        [25]   // Subsurface Cutter Alarm Tone Generation Counter
        [11]   // TRIM DECK Fault Tracking: Number of Times M2CM12N Drive Faulted
        [12]   // TRIM DECK Fault Tracking: Number of Times M2CM04N Drive Faulted
        [18]   // TRIM DECK Fault Tracking: Number of Times M2CM10S Drive Faulted
        [1]   // TRIM DECK Fault Tracking: Number of Times M2CM02 Drive Faulted
        [19]   // TRIM DECK Fault Tracking: Number of Times M2CM11S Drive Faulted
        [22]   // Debug Counter Number of Times M2CM09 Drive Faulted
        [23]   // Debug Counter Number of Times M2CM10 Drive Faulted
        [30]   // TRIM DECK Fault Tracking: Number of Times M2CM01 Drive is Stopped
   C50 : COUNTER[33];
        [10]   // Conveyor 10 Phantom Caps Generated Counter
        [11]   // Conveyor 11 Phantom Caps Generated Counter
        [12]   // Conveyor 12 Phantom Caps Generated Counter
        [13]   // Conveyor 13 Phantom Caps Generated Counter
        [14]   // Conveyor 14 Phantom Caps Generated Counter
        [15]   // Conveyor 15 Phantom Caps Generated Counter
        [16]   // Conveyor 16 Phantom Caps Generated Counter
        [17]   // Conveyor 17 Phantom Caps Generated Counter
        [18]   // Conveyor 18 Phantom Caps Generated Counter
        [19]   // Conveyor 19 Phantom Caps Generated Counter
        [1]   // Conveyor 1 Phantom Caps Generated Counter
        [20]   // Conveyor 20 Phantom Caps Generated Counter
        [21]   // Conveyor 21 Phantom Caps Generated Counter
        [22]   // Conveyor 22 Phantom Caps Generated Counter
        [23]   // Conveyor 23 Phantom Caps Generated Counter
        [24]   // Conveyor 24 Phantom Caps Generated Counter
        [25]   // Conveyor 25 Phantom Caps Generated Counter
        [26]   // Conveyor 26 Phantom Caps Generated Counter
        [27]   // Conveyor 27 Phantom Caps Generated Counter
        [28]   // Conveyor 28 Phantom Caps Generated Counter
        [29]   // Conveyor 29 Phantom Caps Generated Counter
        [2]   // Conveyor 2 Phantom Caps Generated Counter
        [30]   // Conveyor 30 Phantom Caps Generated Counter
        [31]   // Conveyor 31 Phantom Caps Generated Counter
        [32]   // Conveyor 32 Phantom Caps Generated Counter
        [3]   // Conveyor 3 Phantom Caps Generated Counter
        [4]   // Conveyor 4 Phantom Caps Generated Counter
        [5]   // Conveyor 5 Phantom Caps Generated Counter
        [6]   // Conveyor 6 Phantom Caps Generated Counter
        [7]   // Conveyor 7 Phantom Caps Generated Counter
        [8]   // Conveyor 8 Phantom Caps Generated Counter
        [9]   // Conveyor 9 Phantom Caps Generated Counter
   C61 : COUNTER[33];
        [5]   // Conveyor 5 Glass in Transit Counter
        [6]   // Conveyor 6 Glass in Transit Counter
        [7]   // Conveyor 7 Glass in Transit Counter
        [8]   // Conveyor 8 Glass in Transit Counter
        [9]   // Conveyor 9 Glass in Transit Counter
        [17]   // Conveyor 17 Glass in Transit Counter
        [18]   // Conveyor 18 Glass in Transit Counter
        [19]   // Conveyor 19 Glass in Transit Counter
        [1]   // Conveyor 1 Glass in Transit Counter
        [20]   // Conveyor 20 Glass in Transit Counter
        [21]   // Conveyor 21 Glass in Transit Counter
        [22]   // Conveyor 22 Glass in Transit Counter
        [23]   // Conveyor 23 Glass in Transit Counter
        [24]   // Conveyor 24 Glass in Transit Counter
        [25]   // Conveyor 25 Glass in Transit Counter
        [26]   // Conveyor 26 Glass in Transit Counter
        [27]   // Conveyor 27 Glass in Transit Counter
        [10]   // Conveyor 10 Glass in Transit Counter
        [11]   // Conveyor 11 Glass in Transit Counter
        [12]   // Conveyor 12 Glass in Transit Counter
        [13]   // Conveyor 13 Glass in Transit Counter
        [14]   // Conveyor 14 Glass in Transit Counter
        [15]   // Conveyor 15 Glass in Transit Counter
        [28]   // Conveyor 28 Glass in Transit Counter
        [29]   // Conveyor 29 Glass in Transit Counter
        [2]   // Conveyor 2 Glass in Transit Counter
        [16]   // Conveyor 16 Glass in Transit Counter
        [30]   // Conveyor 30 Glass in Transit Counter
        [31]   // Conveyor 31 Glass in Transit Counter
        [32]   // Conveyor 32 Glass in Transit Counter
        [3]   // Conveyor 3 Glass in Transit Counter
        [4]   // Conveyor 4 Glass in Transit Counter
   CM_AreaStackerToLine_JS1 : CM_AreaStackerToLine; {access Read Only}
   CM_AreaStackerToLine_JS1_Sync : CM_AreaStackerToLine := (dSyncHead := 612195157, xAreaOk := 1, xStackerInUnloaderMode := 1, iPresetNumberPlateOnRack[0] := 30, iPresetNumberPlateOnRack[1] := 30, iActualNumberPlateOnRack[0] := 24, iActualNumberPlateOnRack[1] := 23, dGap_cmm := 25000, dMsgDataSyncFdbk := 230589, dMsgDataSync := 289, dMsgOPTSyncFdbk := 339568305, dMsgOPTSync := 297768899, dSyncTail := 612195157);
        .iPresetNumberPlateOnRack[0]   // RHS
        .iActualNumberPlateOnRack[0]   // RHS
        .iActualNumberPlateOnRack[1]   // LHS
        .iPresetNumberPlateOnRack[1]   // LHS
        .dGap_cmm   // [mm/100]
   CM_AreaStackerToLine_JS2 : CM_AreaStackerToLine; {access Read Only}
   CM_AreaStackerToLine_JS2_Sync : CM_AreaStackerToLine := (dSyncHead := 612195157, xAreaOk := 1, xStackerInUnloaderMode := 1, iPresetNumberPlateOnRack[0] := 30, iPresetNumberPlateOnRack[1] := 30, iActualNumberPlateOnRack[0] := 24, iActualNumberPlateOnRack[1] := 23, dGap_cmm := 25000, dMsgDataSyncFdbk := 230589, dMsgDataSync := 289, dMsgOPTSyncFdbk := 339568305, dMsgOPTSync := 297768899, dSyncTail := 612195157);
        .iPresetNumberPlateOnRack[0]   // RHS
        .iPresetNumberPlateOnRack[1]   // LHS
        .iActualNumberPlateOnRack[0]   // RHS
        .iActualNumberPlateOnRack[1]   // LHS
        .dGap_cmm   // [mm/100]
   CM_ConveyorStackerToLine_JS1 : CM_ConveyorStackerToLine; {access Read Only}
   CM_ConveyorStackerToLine_JS1_Sync : CM_ConveyorStackerToLine := (dSyncHead := 598734532, xCycleOn := 1, xConditionOkForStopCycle := 1, xInitialContionOk := 1, xOutputEnable := 1, xAirMode := 1, dSyncTail := 598734532);
   CM_ConveyorStackerToLine_JS2 : CM_ConveyorStackerToLine; {access Read Only}
   CM_ConveyorStackerToLine_JS2_Sync : CM_ConveyorStackerToLine := (dSyncHead := 598734532, xCycleOn := 1, xConditionOkForStopCycle := 1, xInitialContionOk := 1, xOutputEnable := 1, xAirMode := 1, dSyncTail := 598734532);
   CM_DATA_Snap_Rx : CM_DATA_Z200; {access Read Only}
   CM_DATA_Snap_Rx_TempBuffer : SINT[696]; {access Read Only}
   CM_DATA_Z410_Rx : UDT_PlateData_Convoy; {access Read Only}
   CM_DATA_Z410_Rx_Sync : UDT_PlateData_Convoy; {access Read Only}
   CM_DATA_Z410_Rx_TmpBuffer : SINT[104]; {access Read Only}
   CM_DATA_Z410_Tx : UDT_PlateData_Convoy; {access Read Only}
   CM_DATA_Z410_Tx_MSG : MESSAGE; {access Read Only}
   CM_DATA_Z410_Tx_PH : DINT; {access Read Only}
   CM_DATA_Z410_Tx_TempBuffer : SINT[104]; {access Read Only}
   CM_DATA_Z410_Tx_tmON : TIMER; {access Read Only}
   CM_DATA_Z420_Rx : UDT_PlateData_Convoy; {access Read Only}
   CM_DATA_Z420_Rx_Sync : UDT_PlateData_Convoy; {access Read Only}
   CM_DATA_Z420_Rx_TmpBuffer : SINT[104]; {access Read Only}
   CM_DATA_Z420_Tx : UDT_PlateData_Convoy; {access Read Only}
   CM_DATA_Z420_Tx_MSG : MESSAGE; {access Read Only}
   CM_DATA_Z420_Tx_PH : DINT; {access Read Only}
   CM_DATA_Z420_Tx_TempBuffer : SINT[104]; {access Read Only}
   CM_DATA_Z420_Tx_tmON : TIMER; {access Read Only}
   CM_INPUT_Z200 : CM_INPUT_Z200; {access Read Only}
   CM_INPUT_Z200_Sync : CM_INPUT_Z200; {access Read Only}
   CM_LineToAreaStacker_JS1 : CM_LineToAreaStacker := (dSyncHead := 612195196, xConditionOkForAccessArea := 1, dMsgDataSyncFdbk := 289, dMsgDataSync := 230589, dMsgOPTSyncFdbk := 297768899, dMsgOPTSync := 339568321, dSyncTail := 612195196); {produced}
   CM_LineToAreaStacker_JS2 : CM_LineToAreaStacker := (dSyncHead := 612195196, xConditionOkForAccessArea := 1, dMsgDataSyncFdbk := 289, dMsgDataSync := 230589, dMsgOPTSyncFdbk := 297768899, dMsgOPTSync := 339568321, dSyncTail := 612195196); {produced}
   CM_LineToConveyorStacker_JS1 : CM_LineToConveyorStacker := (dSyncHead := 598734505, xEmergencyOn := 1, xLineCycleOn := 1, xOutputEnable := 1, xReadyToMove := 1, dLineSpeed_dmm_min := 600000, dSyncTail := 598734505); {produced}
   CM_LineToConveyorStacker_JS2 : CM_LineToConveyorStacker := (dSyncHead := 598734505, xEmergencyOn := 1, xLineCycleOn := 1, xOutputEnable := 1, xReadyToMove := 1, dLineSpeed_dmm_min := 600000, dSyncTail := 598734505); {produced}
   CM_OUTPUT_Z200 : CM_OUTPUT_Z200; {access Read Only}
   CNV10_COP_BUFR : ALIAS FOR N31[10];
   CNV10_FLT : ALIAS FOR I[4].9;
   CNV10_FWD : ALIAS FOR O[5].9;
   CNV10_LENGTH : ALIAS FOR N32[10];
   CNV10_LOST : ALIAS FOR C48[10];
   CNV10_PHNTM : ALIAS FOR C50[10];
   CNV10_RES_CAPID : ALIAS FOR N40[10];
   CNV10_RESIN : ALIAS FOR B42[0].10;
   CNV10_RESIN_DEB : ALIAS FOR T47[10];
   CNV10_RESIN_LED : ALIAS FOR B45[0].10;
   CNV10_RESIN_TR : ALIAS FOR B46[0].10;
   CNV10_RESOUT : ALIAS FOR B43[0].10;
   CNV10_REV : ALIAS FOR O[6].9;
   CNV10_RTUNE : ALIAS FOR C49[10];
   CNV10_SS1 : ALIAS FOR O[8].9;
   CNV10_SS2 : ALIAS FOR O[7].9;
   CNV10_T : ALIAS FOR B60[0].10;
   CNV10_T_CNTRS : ALIAS FOR C61[10];
   CNV10_WIN : ALIAS FOR B41[0].10;
   CNV11_COP_BUFR : ALIAS FOR N31[11];
   CNV11_FLT : ALIAS FOR I[4].10;
   CNV11_FWD : ALIAS FOR O[5].10;
   CNV11_LENGTH : ALIAS FOR N32[11];
   CNV11_LOST : ALIAS FOR C48[11];
   CNV11_PHNTM : ALIAS FOR C50[11];
   CNV11_RES_CAPID : ALIAS FOR N40[11];
   CNV11_RESIN : ALIAS FOR B42[0].11;
   CNV11_RESIN_DEB : ALIAS FOR T47[11];
   CNV11_RESIN_LED : ALIAS FOR B45[0].11;
   CNV11_RESIN_TR : ALIAS FOR B46[0].11;
   CNV11_RESOUT : ALIAS FOR B43[0].11;
   CNV11_REV : ALIAS FOR O[6].10;
   CNV11_RTUNE : ALIAS FOR C49[11];
   CNV11_SS1 : ALIAS FOR O[8].10;
   CNV11_SS2 : ALIAS FOR O[7].10;
   CNV11_T : ALIAS FOR B60[0].11;
   CNV11_T_CNTRS : ALIAS FOR C61[11];
   CNV11_WIN : ALIAS FOR B41[0].11;
   CNV12_COP_BUFR : ALIAS FOR N31[12];
   CNV12_FLT : ALIAS FOR I[4].11;
   CNV12_LENGTH : ALIAS FOR N32[12];
   CNV12_LOST : ALIAS FOR C48[12];
   CNV12_PHNTM : ALIAS FOR C50[12];
   CNV12_RES_CAPID : ALIAS FOR N40[12];
   CNV12_RESIN : ALIAS FOR B42[0].12;
   CNV12_RESIN_DEB : ALIAS FOR T47[12];
   CNV12_RESIN_LED : ALIAS FOR B45[0].12;
   CNV12_RESIN_TR : ALIAS FOR B46[0].12;
   CNV12_RESOUT : ALIAS FOR B43[0].12;
   CNV12_REV : ALIAS FOR O[6].11;
   CNV12_RTUNE : ALIAS FOR C49[12];
   CNV12_SS1 : ALIAS FOR O[8].11;
   CNV12_SS2 : ALIAS FOR O[7].11;
   CNV12_T : ALIAS FOR B60[0].12;
   CNV12_T_CNTRS : ALIAS FOR C61[12];
   CNV12_WIN : ALIAS FOR B41[0].12;
   CNV13_COP_BUFR : ALIAS FOR N31[13];
   CNV13_LENGTH : ALIAS FOR N32[13];
   CNV13_LOST : ALIAS FOR C48[13];
   CNV13_PHNTM : ALIAS FOR C50[13];
   CNV13_RES_CAPID : ALIAS FOR N40[13];
   CNV13_RESIN : ALIAS FOR B42[0].13;
   CNV13_RESIN_DEB : ALIAS FOR T47[13];
   CNV13_RESIN_LED : ALIAS FOR B45[0].13;
   CNV13_RESIN_TR : ALIAS FOR B46[0].13;
   CNV13_RESOUT : ALIAS FOR B43[0].13;
   CNV13_RTUNE : ALIAS FOR C49[13];
   CNV13_T : ALIAS FOR B60[0].13;
   CNV13_T_CNTRS : ALIAS FOR C61[13];
   CNV13_WIN : ALIAS FOR B41[0].13;
   CNV14_COP_BUFR : ALIAS FOR N31[14];
   CNV14_LENGTH : ALIAS FOR N32[14];
   CNV14_LOST : ALIAS FOR C48[14];
   CNV14_PHNTM : ALIAS FOR C50[14];
   CNV14_RES_CAPID : ALIAS FOR N40[14];
   CNV14_RESIN : ALIAS FOR B42[0].14;
   CNV14_RESIN_DEB : ALIAS FOR T47[14];
   CNV14_RESIN_LED : ALIAS FOR B45[0].14;
   CNV14_RESIN_TR : ALIAS FOR B46[0].14;
   CNV14_RESOUT : ALIAS FOR B43[0].14;
   CNV14_RTUNE : ALIAS FOR C49[14];
   CNV14_T : ALIAS FOR B60[0].14;
   CNV14_T_CNTRS : ALIAS FOR C61[14];
   CNV14_WIN : ALIAS FOR B41[0].14;
   CNV15_COP_BUFR : ALIAS FOR N31[15];
   CNV15_LENGTH : ALIAS FOR N32[15];
   CNV15_LOST : ALIAS FOR C48[15];
   CNV15_PHNTM : ALIAS FOR C50[15];
   CNV15_RES_CAPID : ALIAS FOR N40[15];
   CNV15_RESIN : ALIAS FOR B42[0].15;
   CNV15_RESIN_DEB : ALIAS FOR T47[15];
   CNV15_RESIN_LED : ALIAS FOR B45[0].15;
   CNV15_RESIN_TR : ALIAS FOR B46[0].15;
   CNV15_RESOUT : ALIAS FOR B43[0].15;
   CNV15_RTUNE : ALIAS FOR C49[15];
   CNV15_T : ALIAS FOR B60[0].15;
   CNV15_T_CNTRS : ALIAS FOR C61[15];
   CNV15_WIN : ALIAS FOR B41[0].15;
   CNV16_COP_BUFR : ALIAS FOR N31[16];
   CNV16_LENGTH : ALIAS FOR N32[16];
   CNV16_LOST : ALIAS FOR C48[16];
   CNV16_PHNTM : ALIAS FOR C50[16];
   CNV16_RES_CAPID : ALIAS FOR N40[16];
   CNV16_RESIN : ALIAS FOR B42[1].0;
   CNV16_RESIN_DEB : ALIAS FOR T47[16];
   CNV16_RESIN_LED : ALIAS FOR B45[1].0;
   CNV16_RESIN_TR : ALIAS FOR B46[1].0;
   CNV16_RESOUT : ALIAS FOR B43[1].0;
   CNV16_RTUNE : ALIAS FOR C49[16];
   CNV16_T : ALIAS FOR B60[1].0;
   CNV16_T_CNTRS : ALIAS FOR C61[16];
   CNV16_WIN : ALIAS FOR B41[1].0;
   CNV17_COP_BUFR : ALIAS FOR N31[17];
   CNV17_LENGTH : ALIAS FOR N32[17];
   CNV17_LOST : ALIAS FOR C48[17];
   CNV17_PHNTM : ALIAS FOR C50[17];
   CNV17_RES_CAPID : ALIAS FOR N40[17];
   CNV17_RESIN : ALIAS FOR B42[1].1;
   CNV17_RESIN_DEB : ALIAS FOR T47[17];
   CNV17_RESIN_LED : ALIAS FOR B45[1].1;
   CNV17_RESIN_TR : ALIAS FOR B46[1].1;
   CNV17_RESOUT : ALIAS FOR B43[1].1;
   CNV17_RTUNE : ALIAS FOR C49[17];
   CNV17_T : ALIAS FOR B60[1].1;
   CNV17_T_CNTRS : ALIAS FOR C61[17];
   CNV17_WIN : ALIAS FOR B41[1].1;
   CNV18_COP_BUFR : ALIAS FOR N31[18];
   CNV18_LENGTH : ALIAS FOR N32[18];
   CNV18_LOST : ALIAS FOR C48[18];
   CNV18_PHNTM : ALIAS FOR C50[18];
   CNV18_RES_CAPID : ALIAS FOR N40[18];
   CNV18_RESIN : ALIAS FOR B42[1].2;
   CNV18_RESIN_DEB : ALIAS FOR T47[18];
   CNV18_RESIN_LED : ALIAS FOR B45[1].2;
   CNV18_RESIN_TR : ALIAS FOR B46[1].2;
   CNV18_RESOUT : ALIAS FOR B43[1].2;
   CNV18_RTUNE : ALIAS FOR C49[18];
   CNV18_T : ALIAS FOR B60[1].2;
   CNV18_T_CNTRS : ALIAS FOR C61[18];
   CNV18_WIN : ALIAS FOR B41[1].2;
   CNV19_COP_BUFR : ALIAS FOR N31[19];
   CNV19_LENGTH : ALIAS FOR N32[19];
   CNV19_LOST : ALIAS FOR C48[19];
   CNV19_PHNTM : ALIAS FOR C50[19];
   CNV19_RES_CAPID : ALIAS FOR N40[19];
   CNV19_RESIN : ALIAS FOR B42[1].3;
   CNV19_RESIN_DEB : ALIAS FOR T47[19];
   CNV19_RESIN_LED : ALIAS FOR B45[1].3;
   CNV19_RESIN_TR : ALIAS FOR B46[1].3;
   CNV19_RESOUT : ALIAS FOR B43[1].3;
   CNV19_RTUNE : ALIAS FOR C49[19];
   CNV19_T : ALIAS FOR B60[1].3;
   CNV19_T_CNTRS : ALIAS FOR C61[19];
   CNV19_WIN : ALIAS FOR B41[1].3;
   CNV1_COP_BUFR : ALIAS FOR N31[1];
   CNV1_FLT : ALIAS FOR I[4].0;
   CNV1_FWD : ALIAS FOR O[5].0;
   CNV1_LENGTH : ALIAS FOR N32[1];
   CNV1_LOST : ALIAS FOR C48[1];
   CNV1_PHNTM : ALIAS FOR C50[1];
   CNV1_RES_CAPID : ALIAS FOR N40[1];
   CNV1_RESIN : ALIAS FOR B42[0].1;
   CNV1_RESIN_DEB : ALIAS FOR T47[1];
   CNV1_RESIN_LED : ALIAS FOR B45[0].1;
   CNV1_RESIN_TR : ALIAS FOR B46[0].1;
   CNV1_RESOUT : ALIAS FOR B43[0].1;
   CNV1_REV : ALIAS FOR O[6].0;
   CNV1_RTUNE : ALIAS FOR C49[1];
   CNV1_SS1 : ALIAS FOR O[8].0;
   CNV1_SS2 : ALIAS FOR O[7].0;
   CNV1_T : ALIAS FOR B60[0].1;
   CNV1_T_CNTRS : ALIAS FOR C61[1];
   CNV1_WIN : ALIAS FOR B41[0].1;
   CNV20_COP_BUFR : ALIAS FOR N31[20];
   CNV20_LENGTH : ALIAS FOR N32[20];
   CNV20_LOST : ALIAS FOR C48[20];
   CNV20_PHNTM : ALIAS FOR C50[20];
   CNV20_RES_CAPID : ALIAS FOR N40[20];
   CNV20_RESIN : ALIAS FOR B42[1].4;
   CNV20_RESIN_DEB : ALIAS FOR T47[20];
   CNV20_RESIN_LED : ALIAS FOR B45[1].4;
   CNV20_RESIN_TR : ALIAS FOR B46[1].4;
   CNV20_RESOUT : ALIAS FOR B43[1].4;
   CNV20_RTUNE : ALIAS FOR C49[20];
   CNV20_T : ALIAS FOR B60[1].4;
   CNV20_T_CNTRS : ALIAS FOR C61[20];
   CNV20_WIN : ALIAS FOR B41[1].4;
   CNV21_COP_BUFR : ALIAS FOR N31[21];
   CNV21_LENGTH : ALIAS FOR N32[21];
   CNV21_LOST : ALIAS FOR C48[21];
   CNV21_PHNTM : ALIAS FOR C50[21];
   CNV21_RES_CAPID : ALIAS FOR N40[21];
   CNV21_RESIN : ALIAS FOR B42[1].5;
   CNV21_RESIN_DEB : ALIAS FOR T47[21];
   CNV21_RESIN_LED : ALIAS FOR B45[1].5;
   CNV21_RESIN_TR : ALIAS FOR B46[1].5;
   CNV21_RESOUT : ALIAS FOR B43[1].5;
   CNV21_RTUNE : ALIAS FOR C49[21];
   CNV21_T : ALIAS FOR B60[1].5;
   CNV21_T_CNTRS : ALIAS FOR C61[21];
   CNV21_WIN : ALIAS FOR B41[1].5;
   CNV22_COP_BUFR : ALIAS FOR N31[22];
   CNV22_LENGTH : ALIAS FOR N32[22];
   CNV22_LOST : ALIAS FOR C48[22];
   CNV22_PHNTM : ALIAS FOR C50[22];
   CNV22_RES_CAPID : ALIAS FOR N40[22];
   CNV22_RESIN : ALIAS FOR B42[1].6;
   CNV22_RESIN_DEB : ALIAS FOR T47[22];
   CNV22_RESIN_LED : ALIAS FOR B45[1].6;
   CNV22_RESIN_TR : ALIAS FOR B46[1].6;
   CNV22_RESOUT : ALIAS FOR B43[1].6;
   CNV22_RTUNE : ALIAS FOR C49[22];
   CNV22_T : ALIAS FOR B60[1].6;
   CNV22_T_CNTRS : ALIAS FOR C61[22];
   CNV22_WIN : ALIAS FOR B41[1].6;
   CNV23_COP_BUFR : ALIAS FOR N31[23];
   CNV23_LENGTH : ALIAS FOR N32[23];
   CNV23_LOST : ALIAS FOR C48[23];
   CNV23_PHNTM : ALIAS FOR C50[23];
   CNV23_RES_CAPID : ALIAS FOR N40[23];
   CNV23_RESIN : ALIAS FOR B42[1].7;
   CNV23_RESIN_DEB : ALIAS FOR T47[23];
   CNV23_RESIN_LED : ALIAS FOR B45[1].7;
   CNV23_RESIN_TR : ALIAS FOR B46[1].7;
   CNV23_RESOUT : ALIAS FOR B43[1].7;
   CNV23_RTUNE : ALIAS FOR C49[23];
   CNV23_T : ALIAS FOR B60[1].7;
   CNV23_T_CNTRS : ALIAS FOR C61[23];
   CNV23_WIN : ALIAS FOR B41[1].7;
   CNV24_COP_BUFR : ALIAS FOR N31[24];
   CNV24_LENGTH : ALIAS FOR N32[24];
   CNV24_LOST : ALIAS FOR C48[24];
   CNV24_PHNTM : ALIAS FOR C50[24];
   CNV24_RES_CAPID : ALIAS FOR N40[24];
   CNV24_RESIN : ALIAS FOR B42[1].8;
   CNV24_RESIN_DEB : ALIAS FOR T47[24];
   CNV24_RESIN_LED : ALIAS FOR B45[1].8;
   CNV24_RESIN_TR : ALIAS FOR B46[1].8;
   CNV24_RESOUT : ALIAS FOR B43[1].8;
   CNV24_RTUNE : ALIAS FOR C49[24];
   CNV24_T : ALIAS FOR B60[1].8;
   CNV24_T_CNTRS : ALIAS FOR C61[24];
   CNV24_WIN : ALIAS FOR B41[1].8;
   CNV25_COP_BUFR : ALIAS FOR N31[25];
   CNV25_LENGTH : ALIAS FOR N32[25];
   CNV25_LOST : ALIAS FOR C48[25];
   CNV25_PHNTM : ALIAS FOR C50[25];
   CNV25_RES_CAPID : ALIAS FOR N40[25];
   CNV25_RESIN : ALIAS FOR B42[1].9;
   CNV25_RESIN_DEB : ALIAS FOR T47[25];
   CNV25_RESIN_LED : ALIAS FOR B45[1].9;
   CNV25_RESIN_TR : ALIAS FOR B46[1].9;
   CNV25_RESOUT : ALIAS FOR B43[1].9;
   CNV25_RTUNE : ALIAS FOR C49[25];
   CNV25_T : ALIAS FOR B60[1].9;
   CNV25_T_CNTRS : ALIAS FOR C61[25];
   CNV25_WIN : ALIAS FOR B41[1].9;
   CNV26_COP_BUFR : ALIAS FOR N31[26];
   CNV26_LENGTH : ALIAS FOR N32[26];
   CNV26_LOST : ALIAS FOR C48[26];
   CNV26_PHNTM : ALIAS FOR C50[26];
   CNV26_RES_CAPID : ALIAS FOR N40[26];
   CNV26_RESIN : ALIAS FOR B42[1].10;
   CNV26_RESIN_DEB : ALIAS FOR T47[26];
   CNV26_RESIN_LED : ALIAS FOR B45[1].10;
   CNV26_RESIN_TR : ALIAS FOR B46[1].10;
   CNV26_RESOUT : ALIAS FOR B43[1].10;
   CNV26_RTUNE : ALIAS FOR C49[26];
   CNV26_T : ALIAS FOR B60[1].10;
   CNV26_T_CNTRS : ALIAS FOR C61[26];
   CNV26_WIN : ALIAS FOR B41[1].10;
   CNV27_COP_BUFR : ALIAS FOR N31[27];
   CNV27_LENGTH : ALIAS FOR N32[27];
   CNV27_LOST : ALIAS FOR C48[27];
   CNV27_PHNTM : ALIAS FOR C50[27];
   CNV27_RES_CAPID : ALIAS FOR N40[27];
   CNV27_RESIN : ALIAS FOR B42[1].11;
   CNV27_RESIN_DEB : ALIAS FOR T47[27];
   CNV27_RESIN_LED : ALIAS FOR B45[1].11;
   CNV27_RESIN_TR : ALIAS FOR B46[1].11;
   CNV27_RESOUT : ALIAS FOR B43[1].11;
   CNV27_RTUNE : ALIAS FOR C49[27];
   CNV27_T : ALIAS FOR B60[1].11;
   CNV27_T_CNTRS : ALIAS FOR C61[27];
   CNV27_WIN : ALIAS FOR B41[1].11;
   CNV28_COP_BUFR : ALIAS FOR N31[28];
   CNV28_LENGTH : ALIAS FOR N32[28];
   CNV28_LOST : ALIAS FOR C48[28];
   CNV28_PHNTM : ALIAS FOR C50[28];
   CNV28_RES_CAPID : ALIAS FOR N40[28];
   CNV28_RESIN : ALIAS FOR B42[1].12;
   CNV28_RESIN_DEB : ALIAS FOR T47[28];
   CNV28_RESIN_LED : ALIAS FOR B45[1].12;
   CNV28_RESIN_TR : ALIAS FOR B46[1].12;
   CNV28_RESOUT : ALIAS FOR B43[1].12;
   CNV28_RTUNE : ALIAS FOR C49[28];
   CNV28_T : ALIAS FOR B60[1].12;
   CNV28_T_CNTRS : ALIAS FOR C61[28];
   CNV28_WIN : ALIAS FOR B41[1].12;
   CNV29_COP_BUFR : ALIAS FOR N31[29];
   CNV29_LENGTH : ALIAS FOR N32[29];
   CNV29_LOST : ALIAS FOR C48[29];
   CNV29_PHNTM : ALIAS FOR C50[29];
   CNV29_RES_CAPID : ALIAS FOR N40[29];
   CNV29_RESIN : ALIAS FOR B42[1].13;
   CNV29_RESIN_DEB : ALIAS FOR T47[29];
   CNV29_RESIN_LED : ALIAS FOR B45[1].13;
   CNV29_RESIN_TR : ALIAS FOR B46[1].13;
   CNV29_RESOUT : ALIAS FOR B43[1].13;
   CNV29_RTUNE : ALIAS FOR C49[29];
   CNV29_T : ALIAS FOR B60[1].13;
   CNV29_T_CNTRS : ALIAS FOR C61[29];
   CNV29_WIN : ALIAS FOR B41[1].13;
   CNV2_COP_BUFR : ALIAS FOR N31[2];
   CNV2_FLT : ALIAS FOR I[4].1;
   CNV2_FWD : ALIAS FOR O[5].1;
   CNV2_LENGTH : ALIAS FOR N32[2];
   CNV2_LOST : ALIAS FOR C48[2];
   CNV2_PHNTM : ALIAS FOR C50[2];
   CNV2_RES_CAPID : ALIAS FOR N40[2];
   CNV2_RESIN : ALIAS FOR B42[0].2;
   CNV2_RESIN_DEB : ALIAS FOR T47[2];
   CNV2_RESIN_LED : ALIAS FOR B45[0].2;
   CNV2_RESIN_TR : ALIAS FOR B46[0].2;
   CNV2_RESOUT : ALIAS FOR B43[0].2;
   CNV2_REV : ALIAS FOR O[6].1;
   CNV2_RTUNE : ALIAS FOR C49[2];
   CNV2_SS1 : ALIAS FOR O[8].1;
   CNV2_SS2 : ALIAS FOR O[7].1;
   CNV2_T : ALIAS FOR B60[0].2;
   CNV2_T_CNTRS : ALIAS FOR C61[2];
   CNV2_WIN : ALIAS FOR B41[0].2;
   CNV30_COP_BUFR : ALIAS FOR N31[30];
   CNV30_LENGTH : ALIAS FOR N32[30];
   CNV30_LOST : ALIAS FOR C48[30];
   CNV30_PHNTM : ALIAS FOR C50[30];
   CNV30_RES_CAPID : ALIAS FOR N40[30];
   CNV30_RESIN : ALIAS FOR B42[1].14;
   CNV30_RESIN_DEB : ALIAS FOR T47[30];
   CNV30_RESIN_LED : ALIAS FOR B45[1].14;
   CNV30_RESIN_TR : ALIAS FOR B46[1].14;
   CNV30_RESOUT : ALIAS FOR B43[1].14;
   CNV30_RTUNE : ALIAS FOR C49[30];
   CNV30_T : ALIAS FOR B60[1].14;
   CNV30_T_CNTRS : ALIAS FOR C61[30];
   CNV30_WIN : ALIAS FOR B41[1].14;
   CNV31_COP_BUFR : ALIAS FOR N31[31];
   CNV31_LENGTH : ALIAS FOR N32[31];
   CNV31_LOST : ALIAS FOR C48[31];
   CNV31_PHNTM : ALIAS FOR C50[31];
   CNV31_RES_CAPID : ALIAS FOR N40[31];
   CNV31_RESIN : ALIAS FOR B42[1].15;
   CNV31_RESIN_DEB : ALIAS FOR T47[31];
   CNV31_RESIN_LED : ALIAS FOR B45[1].15;
   CNV31_RESIN_TR : ALIAS FOR B46[1].15;
   CNV31_RESOUT : ALIAS FOR B43[1].15;
   CNV31_RTUNE : ALIAS FOR C49[31];
   CNV31_T : ALIAS FOR B60[1].15;
   CNV31_T_CNTRS : ALIAS FOR C61[31];
   CNV31_WIN : ALIAS FOR B41[1].15;
   CNV32_COP_BUFR : ALIAS FOR N31[32];
   CNV32_LENGTH : ALIAS FOR N32[32];
   CNV32_LOST : ALIAS FOR C48[32];
   CNV32_PHNTM : ALIAS FOR C50[32];
   CNV32_RESIN : ALIAS FOR B42[2].0;
   CNV32_RESIN_LED : ALIAS FOR B45[2].0;
   CNV32_RESIN_TR : ALIAS FOR B46[2].0;
   CNV32_RESOUT : ALIAS FOR B43[2].0;
   CNV32_RTUNE : ALIAS FOR C49[32];
   CNV32_T : ALIAS FOR B60[2].0;
   CNV32_T_CNTRS : ALIAS FOR C61[32];
   CNV32_WIN : ALIAS FOR B41[2].0;
   CNV3_COP_BUFR : ALIAS FOR N31[3];
   CNV3_FLT : ALIAS FOR I[4].2;
   CNV3_FWD : ALIAS FOR O[5].2;
   CNV3_LENGTH : ALIAS FOR N32[3];
   CNV3_LOST : ALIAS FOR C48[3];
   CNV3_PHNTM : ALIAS FOR C50[3];
   CNV3_RES_CAPID : ALIAS FOR N40[3];
   CNV3_RESIN : ALIAS FOR B42[0].3;
   CNV3_RESIN_DEB : ALIAS FOR T47[3];
   CNV3_RESIN_LED : ALIAS FOR B45[0].3;
   CNV3_RESIN_TR : ALIAS FOR B46[0].3;
   CNV3_RESOUT : ALIAS FOR B43[0].3;
   CNV3_REV : ALIAS FOR O[6].2;
   CNV3_RTUNE : ALIAS FOR C49[3];
   CNV3_SS1 : ALIAS FOR O[8].2;
   CNV3_SS2 : ALIAS FOR O[7].2;
   CNV3_T : ALIAS FOR B60[0].3;
   CNV3_T_CNTRS : ALIAS FOR C61[3];
   CNV3_WIN : ALIAS FOR B41[0].3;
   CNV4_COP_BUFR : ALIAS FOR N31[4];
   CNV4_FLT : ALIAS FOR I[4].3;
   CNV4_FWD : ALIAS FOR O[5].3;
   CNV4_LENGTH : ALIAS FOR N32[4];
   CNV4_LOST : ALIAS FOR C48[4];
   CNV4_PHNTM : ALIAS FOR C50[4];
   CNV4_RES_CAPID : ALIAS FOR N40[4];
   CNV4_RESIN : ALIAS FOR B42[0].4;
   CNV4_RESIN_DEB : ALIAS FOR T47[4];
   CNV4_RESIN_LED : ALIAS FOR B45[0].4;
   CNV4_RESIN_TR : ALIAS FOR B46[0].4;
   CNV4_RESOUT : ALIAS FOR B43[0].4;
   CNV4_REV : ALIAS FOR O[6].3;
   CNV4_RTUNE : ALIAS FOR C49[4];
   CNV4_SS1 : ALIAS FOR O[8].3;
   CNV4_SS2 : ALIAS FOR O[7].3;
   CNV4_T : ALIAS FOR B60[0].4;
   CNV4_T_CNTRS : ALIAS FOR C61[4];
   CNV4_WIN : ALIAS FOR B41[0].4;
   CNV5_COP_BUFR : ALIAS FOR N31[5];
   CNV5_FLT : ALIAS FOR I[4].4;
   CNV5_FWD : ALIAS FOR O[5].4;
   CNV5_LENGTH : ALIAS FOR N32[5];
   CNV5_LOST : ALIAS FOR C48[5];
   CNV5_PHNTM : ALIAS FOR C50[5];
   CNV5_RES_CAPID : ALIAS FOR N40[5];
   CNV5_RESIN : ALIAS FOR B42[0].5;
   CNV5_RESIN_DEB : ALIAS FOR T47[5];
   CNV5_RESIN_LED : ALIAS FOR B45[0].5;
   CNV5_RESIN_TR : ALIAS FOR B46[0].5;
   CNV5_RESOUT : ALIAS FOR B43[0].5;
   CNV5_REV : ALIAS FOR O[6].4;
   CNV5_RTUNE : ALIAS FOR C49[5];
   CNV5_SS1 : ALIAS FOR O[8].4;
   CNV5_SS2 : ALIAS FOR O[7].4;
   CNV5_T : ALIAS FOR B60[0].5;
   CNV5_T_CNTRS : ALIAS FOR C61[5];
   CNV5_WIN : ALIAS FOR B41[0].5;
   CNV6_COP_BUFR : ALIAS FOR N31[6];
   CNV6_FLT : ALIAS FOR I[4].5;
   CNV6_FWD : ALIAS FOR O[5].5;
   CNV6_LENGTH : ALIAS FOR N32[6];
   CNV6_LOST : ALIAS FOR C48[6];
   CNV6_PHNTM : ALIAS FOR C50[6];
   CNV6_RES_CAPID : ALIAS FOR N40[6];
   CNV6_RESIN : ALIAS FOR B42[0].6;
   CNV6_RESIN_DEB : ALIAS FOR T47[6];
   CNV6_RESIN_LED : ALIAS FOR B45[0].6;
   CNV6_RESIN_TR : ALIAS FOR B46[0].6;
   CNV6_RESOUT : ALIAS FOR B43[0].6;
   CNV6_REV : ALIAS FOR O[6].5;
   CNV6_RTUNE : ALIAS FOR C49[6];
   CNV6_SS1 : ALIAS FOR O[8].5;
   CNV6_SS2 : ALIAS FOR O[7].5;
   CNV6_T : ALIAS FOR B60[0].6;
   CNV6_T_CNTRS : ALIAS FOR C61[6];
   CNV6_WIN : ALIAS FOR B41[0].6;
   CNV7_COP_BUFR : ALIAS FOR N31[7];
   CNV7_FLT : ALIAS FOR I[4].6;
   CNV7_FWD : ALIAS FOR O[5].6;
   CNV7_LENGTH : ALIAS FOR N32[7];
   CNV7_LOST : ALIAS FOR C48[7];
   CNV7_PHNTM : ALIAS FOR C50[7];
   CNV7_RES_CAPID : ALIAS FOR N40[7];
   CNV7_RESIN : ALIAS FOR B42[0].7;
   CNV7_RESIN_DEB : ALIAS FOR T47[7];
   CNV7_RESIN_LED : ALIAS FOR B45[0].7;
   CNV7_RESIN_TR : ALIAS FOR B46[0].7;
   CNV7_RESOUT : ALIAS FOR B43[0].7;
   CNV7_REV : ALIAS FOR O[6].6;
   CNV7_RTUNE : ALIAS FOR C49[7];
   CNV7_SS1 : ALIAS FOR O[8].6;
   CNV7_SS2 : ALIAS FOR O[7].6;
   CNV7_T : ALIAS FOR B60[0].7;
   CNV7_T_CNTRS : ALIAS FOR C61[7];
   CNV7_WIN : ALIAS FOR B41[0].7;
   CNV8_COP_BUFR : ALIAS FOR N31[8];
   CNV8_FLT : ALIAS FOR I[4].7;
   CNV8_FWD : ALIAS FOR O[5].7;
   CNV8_LENGTH : ALIAS FOR N32[8];
   CNV8_LOST : ALIAS FOR C48[8];
   CNV8_PHNTM : ALIAS FOR C50[8];
   CNV8_RES_CAPID : ALIAS FOR N40[8];
   CNV8_RES_CAPID1 : ALIAS FOR N40[8];
   CNV8_RESIN : ALIAS FOR B42[0].8;
   CNV8_RESIN_DEB : ALIAS FOR T47[8];
   CNV8_RESIN_LED : ALIAS FOR B45[0].8;
   CNV8_RESIN_TR : ALIAS FOR B46[0].8;
   CNV8_RESOUT : ALIAS FOR B43[0].8;
   CNV8_REV : ALIAS FOR O[6].7;
   CNV8_RTUNE : ALIAS FOR C49[8];
   CNV8_SS1 : ALIAS FOR O[8].7;
   CNV8_SS2 : ALIAS FOR O[7].7;
   CNV8_T : ALIAS FOR B60[0].8;
   CNV8_T_CNTRS : ALIAS FOR C61[8];
   CNV8_WIN : ALIAS FOR B41[0].8;
   CNV9_COP_BUFR : ALIAS FOR N31[9];
   CNV9_FLT : ALIAS FOR I[4].8;
   CNV9_FWD : ALIAS FOR O[21].8;
   CNV9_FWD1 : ALIAS FOR O[5].8;
   CNV9_LENGTH : ALIAS FOR N32[9];
   CNV9_LOST : ALIAS FOR C48[9];
   CNV9_PHNTM : ALIAS FOR C50[9];
   CNV9_RES_CAPID : ALIAS FOR N40[9];
   CNV9_RESIN : ALIAS FOR B42[0].9;
   CNV9_RESIN_DEB : ALIAS FOR T47[9];
   CNV9_RESIN_LED : ALIAS FOR B45[0].9;
   CNV9_RESIN_TR : ALIAS FOR B46[0].9;
   CNV9_RESOUT : ALIAS FOR B43[0].9;
   CNV9_REV : ALIAS FOR O[6].8;
   CNV9_RTUNE : ALIAS FOR C49[9];
   CNV9_SS1 : ALIAS FOR O[8].8;
   CNV9_SS2 : ALIAS FOR O[7].8;
   CNV9_T : ALIAS FOR B60[0].9;
   CNV9_T_CNTRS : ALIAS FOR C61[9];
   CNV9_WIN : ALIAS FOR B41[0].9;
   COMMAND_FREQ : ALIAS FOR N7[10];
   CONST_dDest_Cullet : DINT; {access Read Only}
   CONST_dDest_Stk : DINT; {access Read Only}
   Const_Empty_Data : UDT_Convoy_SL;
   CONST_rgdDestMask : DINT[32] := ([0] := 16#0000_0001, [1] := 16#0000_0002, [2] := 16#0000_0004, [3] := 16#0000_0008, [4] := 16#0000_0010, [24] := 16#0100_0000, [29] := 16#2000_0000); {constant, access None}   // Destination Mask
        [0]   // Side leg 1 - ATJS - M410
        [1]   // Side leg 1A - ATJS - M420
        [24]   // Generic cullet
        [29]   // Quality #1 - M352
        [4]   // Side leg 4
        [3]   // Side leg 3
        [30]   // Quality #2 - M353
        [2]   // Side leg 2 - Hager Stacker - M510
        [5]   // Side leg 5
        [6]   // End Line Stacker
        [31]   // Quality #3 - End line
   CONST_tAux : AUX_COSTANTS := (dM302SpeedUpMinGapInConvoy_cmm := 15000, dM310_PopUpCycleTime_s[0] := 8, dM310_PopUpCycleTime_s[1] := 8, dM315_PopUpCycleTime_s[0] := 8, dM315_PopUpCycleTime_s[1] := 8); {access Read Only}
   CONST_tPlant : UDT_PLANT_CONSTANTS := (dPLC_ID := 1, dOP_Side := 1, dZ1ConveyorNumber := 29, dZ1TotalLength_cmm := 5395000, dTrimDeckNumber := 6, dTrimWheelsNumber := 12, dTrackWindows_cmm := 12500, dMaxScanSpace_cmm := 17500, rgdAccDecRamps[0] := 1.25, rgdAccDecRamps[1] := 1.2, rgdAccDecRamps[2] := 2.19, rgdAccDecRamps[3] := 0.7, dMaxLineSpeed_mm_min := 84000, dMinLineSpeed_mm_min := 7000, dMaxLineSnapSpeed_mm_min := 54000, dMinLineSnapSpeed_mm_min := 7000, dMaxLehrSpeed_mm_min := 22500, dMinLehrSpeed_mm_min := 2330, rMaxSpeedRatio := 4.0, rMinSpeedRatio := 1.5, rMaxSpeedSnapRatio := 6.0, rMinSpeedSnapRatio := 2.5, dZ1CleaningSpeed_mm_min := 20000, dMaxNumPlates := 40, dMaxNumHeadTail := 1000, rgdLiteLimits_cmm[0] := 62000, rgdLiteLimits_cmm[1] := 610000, rgdLiteLimits_cmm[2] := 62000, rgdLiteLimits_cmm[3] := 610000, rgdLiteLimits_cmm[4] := 420000, rgdLiteLimits_cmm[5] := 610000, rgdLiteLimits_cmm[6] := 62000, rgdLiteLimits_cmm[7] := 366000, rgdLiteLimits_cmm[8] := 62000, rgdLiteLimits_cmm[9] := 280000, rgdLiteLimits_cmm[10] := 46000, rgdLiteLimits_cmm[11] := 366000, rgdLiteLimits_cmm[12] := 46000, rgdLiteLimits_cmm[13] := 400000, rgdLiteLimits_cmm[14] := 260000, rgdLiteLimits_cmm[15] := 366000, rgdLiteLimits_cmm[16] := 46000, rgdLiteLimits_cmm[17] := 366000, rgdLiteLimits_cmm[18] := 46000, rgdLiteLimits_cmm[19] := 280000, rgdCapLimits_cmm[0] := 7, rgdCapLimits_cmm[1] := 46000, rgdCapLimits_cmm[2] := 368000, rgdConvoyLimits_cmm[0] := 4, rgdConvoyLimits_cmm[1] := 130000, rgdConvoyLimits_cmm[2] := 360000, rgdConvoyLimits_cmm[3] := 62000, rgdConvoyLimits_cmm[4] := 165000, rgdRibbonLimits_cmm[0] := 285000, rgdRibbonLimits_cmm[1] := 400000, rgdRibbonLimits_cmm[2] := 260000, rgdRibbonLimits_cmm[3] := 368000, rgdWanderLimits[0] := -25000, rgdWanderLimits[1] := 25000, dNumOfConveyors := 29,
        dNumCapsConveyor := 10, dNumCapsMaxConvoy := 2, dNumLitesMaxCap := 7, dNumPlateSearch := 5, dNumOfUnloadDestinations := 4); {constant, access None}
        .rgdCapLimits_cmm[0]   // Max number of lites in cap
        .rgdCapLimits_cmm[1]   // Width Min [mm/100]
        .rgdCapLimits_cmm[2]   // Width Max [mm/100]
        .rgdLiteLimits_cmm[0]   // Length Min (to cullet) [mm/100]
        .rgdLiteLimits_cmm[10]   // Width Min (to cullet) [mm/100]
        .rgdLiteLimits_cmm[11]   // Width Max (to cullet) [mm/100]
        .rgdLiteLimits_cmm[12]   // Width Min (to quality) [mm/100]
        .rgdLiteLimits_cmm[13]   // Width Max (to quality) [mm/100]
        .rgdLiteLimits_cmm[14]   // Width Min JS [mm/100]
        .rgdLiteLimits_cmm[15]   // Width Max JS [mm/100]
        .rgdLiteLimits_cmm[16]   // Width Min LES [mm/100]
        .rgdLiteLimits_cmm[17]   // Width Max LES [mm/100]
        .rgdLiteLimits_cmm[18]   // Width Min SSS [mm/100]
        .rgdLiteLimits_cmm[19]   // Width Max SSS [mm/100]
        .rgdLiteLimits_cmm[1]   // Length Max (to cullet) [mm/100]
        .rgdLiteLimits_cmm[2]   // Length Min (to quality) [mm/100]
        .rgdLiteLimits_cmm[3]   // Length Max (to quality) [mm/100]
        .rgdLiteLimits_cmm[4]   // Length Min JS [mm/100]
        .rgdLiteLimits_cmm[5]   // Length Max JS [mm/100]
        .rgdLiteLimits_cmm[6]   // Length Min LES [mm/100]
        .rgdLiteLimits_cmm[7]   // Length Max LES [mm/100]
        .rgdLiteLimits_cmm[8]   // Length Min SSS [mm/100]
        .rgdLiteLimits_cmm[9]   // Length Max SSS [mm/100]
        .rgdRibbonLimits_cmm[0]   // Gross width Min [mm/100]
        .rgdRibbonLimits_cmm[1]   // Gross width Max [mm/100]
        .rgdRibbonLimits_cmm[2]   // Net width Min [mm/100]
        .rgdRibbonLimits_cmm[3]   // Net width Max [mm/100]
        .rgdWanderLimits[0]   // Min [mm/100]
        .rgdWanderLimits[1]   // Max [mm/100]
        .rgdConvoyLimits_cmm[0]   // Max number cap in convoy
        .rgdConvoyLimits_cmm[1]   // Length Min [mm/100]
        .rgdConvoyLimits_cmm[2]   // Length Max [mm/100]
        .rgdConvoyLimits_cmm[3]   // Minimum cap length for convoy [mm/100]
        .rgdConvoyLimits_cmm[4]   // Maximum cap length for convoy [mm/100]
        .rgdAccDecRamps[0]   // Speed limit for lower ramps [mm/min]
        .rgdAccDecRamps[1]   // Acceleration / Deceleration with lower speed [m/s2]
        .rgdAccDecRamps[2]   // Speed limit for highest ramps [mm/min]
        .rgdAccDecRamps[3]   // Acceleration / Deceleration with highest speed [m/s2]
   CONV10_MS_ACCUM : ALIAS FOR N30[10];
   CONV11_MS_ACCUM : ALIAS FOR N30[11];
   CONV12_MS_ACCUM : ALIAS FOR N30[12];
   CONV13_MS_ACCUM : ALIAS FOR N30[13];
   CONV14_MS_ACCUM : ALIAS FOR N30[14];
   CONV15_MS_ACCUM : ALIAS FOR N30[15];
   CONV16_MS_ACCUM : ALIAS FOR N30[16];
   CONV17_MS_ACCUM : ALIAS FOR N30[17];
   CONV18_MS_ACCUM : ALIAS FOR N30[18];
   CONV19_MS_ACCUM : ALIAS FOR N30[19];
   CONV1_MS_ACCUM : ALIAS FOR N30[1];
   CONV20_MS_ACCUM : ALIAS FOR N30[20];
   CONV21_MS_ACCUM : ALIAS FOR N30[21];
   CONV22_MS_ACCUM : ALIAS FOR N30[22];
   CONV23_MS_ACCUM : ALIAS FOR N30[23];
   CONV24_MS_ACCUM : ALIAS FOR N30[24];
   CONV25_MS_ACCUM : ALIAS FOR N30[25];
   CONV26_MS_ACCUM : ALIAS FOR N30[26];
   CONV27_MS_ACCUM : ALIAS FOR N30[27];
   CONV28_MS_ACCUM : ALIAS FOR N30[28];
   CONV29_MS_ACCUM : ALIAS FOR N30[29];
   CONV2_MS_ACCUM : ALIAS FOR N30[2];
   CONV30_MS_ACCUM : ALIAS FOR N30[30];
   CONV31_MS_ACCUM : ALIAS FOR N30[31];
   CONV3_MS_ACCUM : ALIAS FOR N30[3];
   CONV4_MS_ACCUM : ALIAS FOR N30[4];
   CONV5_MS_ACCUM : ALIAS FOR N30[5];
   CONV6_MS_ACCUM : ALIAS FOR N30[6];
   CONV7_MS_ACCUM : ALIAS FOR N30[7];
   CONV8_MS_ACCUM : ALIAS FOR N30[8];
   CONV9_MS_ACCUM : ALIAS FOR N30[9];
   Convoy_SL_DATA_NULL : UDT_Convoy_SL; {access Read Only}
   CRUSH_ALL_ON : ALIAS FOR B3[0].0;
   DROP_NO1_CRSH : ALIAS FOR I[73].12;
   DRV_STOP_DEB : ALIAS FOR T4[30].DN;
   ECL_HLD_AUTO : ALIAS FOR N14[240].2;
   ECL_HLD_AUTO_N : ALIAS FOR I[36].14;
   ECL_HLD_AUTO_S : ALIAS FOR I[80].14;
   ECL_HLD_UP : ALIAS FOR N14[240].3;
   ECL_HLD_UP_N : ALIAS FOR I[36].15;
   ECL_HLD_UP_S : ALIAS FOR I[80].15;
   F34 : REAL[2] := ([0] := 50.0, [1] := 0.04);
   F8 : REAL[51];
   F96 : REAL[31] := ([0] := 471.5);
        [21]   // LEHR SPEED Table of Lehr speed Samples over Ten seconds
        [11]   // LEHR SPEED Information Received from Reliance Capping system
        [10]   // LEHR SPEED Information Received from Reliance AutoMax
        [5]   // LEHR SPEED Current Lehr Lower Limit
        [20]   // LEHR SPEED Table of Speed samples Over last ten Seconds
        [0]   // LEHR SPEED Current lehr Speed used Setting Speed of drives
        [6]   // LEHR SPEED Current Lehr Speed upper Limit
        [1]   // LEHR SPEED Average lehr Speed Calculated from Sample table
   FAST_BLINK : ALIAS FOR T4[2];
   FL_HLD_AUTO : ALIAS FOR N14[240].0;
   FL_HLD_AUTO_N : ALIAS FOR I[36].12;
   FL_HLD_AUTO_S : ALIAS FOR I[80].12;
   FL_HLD_UP : ALIAS FOR N14[240].1;
   FL_HLD_UP_N : ALIAS FOR I[36].13;
   FL_HLD_UP_S : ALIAS FOR I[80].13;
   GP_AccessArea_M311S : GP_AccessArea; {access Read Only}
   GP_AccessArea_M311S_STC : GP_AccessArea_STC; {access Read Only}
   GP_AccessArea_M316S : GP_AccessArea;
   GP_AccessArea_M316S_STC : GP_AccessArea_STC; {access Read Only}
   GP_AccTimeForGap : GP_AccTimeForGap; {access Read Only}
   GP_CheckIdPlatePresent : GP_CheckIdPlatePresent; {access Read Only}
   GP_CompactConvoy : GP_CompactConvoy; {access Read Only}
   GP_ConversionXY : GP_ConversionXY; {access Read Only}
   GP_ConvertDataFromStacker : GP_ConvertDataFromStacker; {access Read Only}
   GP_ConvertDataToStacker : GP_ConvertDataToStacker; {access Read Only}
   GP_InvertCapxLite : GP_InvertCapxLite; {access Read Only}
   GP_M311A : GP_Rotator; {access Read Only}
   GP_M316A : GP_Rotator; {access Read Only}
   GP_NetDiag : GP_NetworkDiag;
   GP_OB_InitializeDiag : GP_OB_Initialize;
   GP_OB_InitializeDiag_STC : GP_OB_Initialize_STC;
   GP_OB_InitializeMain : GP_OB_Initialize; {access Read Only}
   GP_OB_InitializeMain_STC : GP_OB_Initialize_STC; {access Read Only}
   GP_PlateYPosition : GP_PlateYPosition; {access Read Only}
   GP_PosWindow : GP_PosWindow; {access Read Only}
   GP_RampManagement : GP_RampManagement; {access Read Only}
   GP_RampSpace : GP_RampSpace; {access Read Only}
   GP_ScadaPlate : GP_ScadaPlate; {access Read Only}
   Gp_SpaceConvUtilities_V1 : GP_SpaceConvUtilities_V1; {access Read Only}
   GP_TrackingAddCap : GP_TrackingAddCap; {access Read Only}
   GP_TrackingFiring : GP_TrackingFiring; {access Read Only}
   GP_TrackingFiringForConvoy : GP_TrackingFiringForConvoy; {access Read Only}
   GP_TrackingGetFirstPlateInConveyor : GP_TrackingGetFirstPlateInConveyor; {access Read Only}
   GP_TrackingGetLength : GP_TrackingGetLength; {access Read Only}
   GP_TrackingPresencePlate : GP_TrackingPresencePlate; {access Read Only}
   GP_TrackingSearchPlate : GP_TrackingSearchPlate; {access Read Only}
   GP_TrackingValidateIndex : GP_TrackingValidateIndex; {access Read Only}
   HMI_Alarm_Presence : BOOL := 1;   // HMI_Alarm_Presence
   HMI_Alarms_0 : BOOL[32] := ([12] := 1, [13] := 1);   // HMI Alarms
   HMI_Alarms_1 : BOOL[32] := ([12] := 1, [13] := 1);   // HMI Alarms
   HMI_Alarms_2 : BOOL[32];   // HMI Alarms
   HMI_Alarms_3 : BOOL[32];   // HMI Alarms
   HMI_Alarms_4 : BOOL[32];   // HMI Alarms
   HMI_Alarms_5 : BOOL[32];   // HMI Alarms
   HMI_Alarms_6 : BOOL[32];   // HMI Alarms
   HMI_Alarms_7 : BOOL[32];   // HMI Alarms
   HMI_Alarms_8 : BOOL[32];   // HMI Alarms
   HMI_Alarms_9 : BOOL[32];   // HMI Alarms
   HMI_Always_ON : BOOL := 1;   // HMI Always ON
   HMI_MAN_CMD_WR : UDT_MAN_CMD_WR; {access Read Only}
   HMI_MOTOR_HMR : UDT_MOTOR_HMR; {access Read Only}
   HMI_Reset_Alarms : BOOL; {access Read Only}
   HOLD_DWN_ECLPS : ALIAS FOR O[38].5;
   HOLD_DWN_FLOAT : ALIAS FOR O[38].4;
   Host_Read : INT[500] := ([2] := 4088, [4] := 4095, [16] := 4095, [22] := 2048, [40] := -1, [41] := -1, [42] := -1, [43] := -1, [44] := 1, [46] := 1, [122] := 4088, [124] := 4095, [136] := 4095, [142] := 2048, [160] := 1, [162] := 1, [164] := 2, [166] := 2, [480] := 10);
   I : INT[128] := ([1] := 2#0000_0011_1111_1100, [2] := 2#0001_0100_1110_1110, [3] := 2#0000_1111_1111_1000, [4] := 2#0000_1111_1111_1111, [17] := 2#0000_0100_1111_1110, [18] := 2#0000_0000_0000_0111, [24] := 2#0101_0000_0111_1001, [26] := 2#0000_0011_1000_0000, [27] := 2#0000_1111_0000_1111, [28] := 2#0000_0011_1000_0000, [29] := 2#0000_1111_0000_1111, [30] := 2#0000_0011_1000_0000, [31] := 2#0000_1111_0000_1111, [53] := 2#0000_0000_0010_0000, [57] := 2#0000_0000_0010_0000, [73] := 2#1010_0000_0000_0000, [84] := 2#0000_0011_1000_0000, [85] := 2#0011_1011_0000_1111, [86] := 2#0000_0011_1000_0000, [87] := 2#0011_1111_0000_1111, [88] := 2#0000_0011_1000_0000, [89] := 2#0011_1111_0000_1111, [90] := 2#0000_0011_1000_0000, [91] := 2#0011_1111_0000_1111, [92] := 2#0000_0011_1000_0000, [93] := 2#0011_1111_0000_1111, [94] := 2#0000_0011_1000_0000, [95] := 2#0011_1111_0000_1111, [96] := 2#0000_0011_1000_0000, [97] := 2#0011_1111_0000_1111, [98] := 2#0000_0011_1000_0000, [99] := 2#0011_1111_0000_1111, [100] := 2#0000_0011_1000_0000, [101] := 2#0011_1011_0000_1111, [102] := 2#0000_0011_1000_0000, [103] := 2#0011_1111_0000_1111, [104] := 2#0000_0011_1000_0000, [105] := 2#0011_1111_0000_1111, [106] := 2#0000_0011_1000_0000, [107] := 2#0011_1111_0000_1111, [108] := 2#0000_0011_1000_0000, [109] := 2#0011_1111_0000_1111, [110] := 2#0000_0011_1000_0000, [111] := 2#0011_1111_0000_1111, [112] := 2#0000_0011_1000_0000, [113] := 2#0011_1111_0000_1111, [114] := 2#0000_0011_1000_0000, [115] := 2#0011_1111_0000_1111, [116] := 2#0000_0011_1000_0000, [117] := 2#0011_1111_0000_1111, [118] := 2#0000_0011_1000_0000, [119] := 2#0011_1111_0000_1111, [121] := 2#0000_0100_1101_0010, [123] := 2#0000_0000_0001_1010, [124] := 2#0000_0101_0010_1000);   // Local Input Updates Input Slot 2
        [56].5   // PANEL TD-CS5S Trim knocker #5 Move DOWN South Selector Sw.
        [76].11   // PANEL KD-CS1S Knurl knocker Move DOWN North Selector Sw.
        [125]   // RELIANCE CAPPER Inputs for Crossbreak (0) And Y-cut Diables
        [32].0   // PANEL KD-CS1N Knurl knocker Move IN South Selector Sw.
        [101].2   // Command direction FW M2CM8S
        [72].0   // BENCHBOARD Trim knocker #1 North Up Selector Sw.
        [72].2   // BENCHBOARD Trim knocker #1 South Up Selector Sw.
        [32].10   // PANEL KD-CS1N Knurl knocker Move UP North Selector Sw.
        [101].8   // Drive at speed M2CM8S
        [103].8   // Drive at speed M2CM8N
        [101].1   // Drive running M2CM8S
        [109].9   // Local control 1 M2CM10S
        [101].4   // Accelerating M2CM8S
        [101].5   // Decelerating M2CM8S
        [16]   // RACK 2 INPUT UPDATES
        [2].9   // VMCC M2 Alarm Reset
        [111].9   // Local control 1 M2CM10N
        [24]   // RACK 3 INPUT UPDATES
        [26]   // RACK 3 INPUT UPDATES
        [64]   // RACK 10 INPUT UPDATES
        [28]   // RACK 3 INPUT UPDATES
        [30]   // RACK 3 INPUT UPDATES
        [101].6   // Drive has an alarm M2CM8S
        [103].11   // Local control 3 M2CM8N
        [105].8   // Drive at speed M2CM9S
        [107].8   // Drive at speed M2CM9N
        [109].1   // Drive running M2CM10S
        [111].1   // Drive running M2CM10N
        [103].1   // Drive running M2CM8N
        [113].9   // Local control 1 M2CM11S
        [103].4   // Accelerating M2CM8N
        [103].5   // Decelerating M2CM8N
        [32]   // RACK 4 INPUT UPDATES
        [68]   // RACK 10 INPUT UPDATES
        [115].9   // Local control 1 M2CM11N
        [101].0   // Drive ready M2CM8S
        [101].12   // Speed reference 1 M2CM8S
        [101].13   // Speed reference 2 M2CM8S
        [101].14   // Speed reference 3 M2CM8S
        [32].5   // PANEL KD-CS1N Knurl knocker Move DOWN South Selector Sw.
        [36]   // RACK 4 INPUT UPDATES
        [40]   // RACK 5 INPUT UPDATES
        [72]   // RACK 11 INPUT UPDATES
        [44]   // RACK 5 INPUT UPDATES
        [48]   // RACK 6 INPUT UPDATES
        [103].6   // Drive has an alarm M2CM8N
        [103].7   // Drive has a fault M2CM8N
        [113].1   // Drive running M2CM11S
        [115].1   // Drive running M2CM11N
        [117].1   // Drive running M2CM12S
        [119].1   // Drive running M2CM12N
        [105].1   // Drive running M2CM9S
        [117].9   // Local control 1 M2CM12S
        [105].4   // Accelerating M2CM9S
        [105].5   // Decelerating M2CM9S
        [50]   // RACK 5 INPUT UPDATES
        [76]   // RACK 11 INPUT UPDATES
        [119].8   // Drive at speed M2CM12N
        [103].0   // Drive ready M2CM8N
        [52]   // RACK 6 INPUT UPDATES
        [54]   // RACK 5 INPUT UPDATES
        [80]   // RACK 12 INPUT UPDATES
        [56]   // RACK 7 INPUT UPDATES
        [60]   // RACK 7 INPUT UPDATES
        [105].10   // Local control 2 M2CM9S
        [105].11   // Local control 3 M2CM9S
        [119].5   // Decelerating M2CM12N
        [17].10   // VMCC TD E-STOP ACTIVE
        [17].5   // VMCC TD E-STOP Power ON
        [29].7   // Drive has a fault M2CM2
        [107].1   // Drive running M2CM9N
        [119].9   // Local control 1 M2CM12N
        [107].4   // Accelerating M2CM9N
        [107].5   // Decelerating M2CM9N
        [70]   // RACK 7 INPUT UPDATES
        [84]   // RACK 12 INPUT UPDATES
        [17].2   // VMCC TD DC Input Power ON
        [105].0   // Drive ready M2CM9S
        [73].8   // BENCHBOARD SPARE
        [73].9   // BENCHBOARD SPARE
        [1].10   // Rockwell Run out Speed up signal M2CM01
        [3].3   // VMCC M2 Speed zone 4 Drive Fault * 2CM04S
        [105].6   // Drive has an alarm M2CM9S
        [125].1   // ROCKWELL CAPPER Input to Disable manual y-cut bar 2
        [24].1   // RELIANCE CAPPING SYSTEM Trim Knocker #1 North Lower wheel
        [32].11   // PANEL KD-CS1N Knurl knocker Move DOWN North Selector Sw.
        [24].2   // RELIANCE CAPPING SYSTEM Trim Knocker #1 South Lower wheel
        [4]   // Word containing Fault bits For trim deck Drives
        [18].1   // VMCC TD Trim deck Drive fault North side
        [123].5   // MB -->> M2 Subsurface Cutters are In Alarm
        [18].2   // VMCC TD Trim deck Drive fault South side
        [24].14   // RELIANCE CAPPING SYSTEM Input Power ON
        [1].0   // Rockwell Run out Speed up signal M2CM2
        [101].10   // Local control 2 M2CM8S
        [109].0   // Drive ready M2CM10S
        [56].15   // PANEL TD-CS5S Reliance Handoff Sensor (Redundant Sensor on South Side)
        [44].12   // Trim Deck PANEL TD-CS3N Crush all OFF Switch
        [73].11   // Reliance BENCHBOARD Crush all ON Switch
        [123].3   // MB -->> M2 No. 1 Crusher Down prox. Made
        [105].2   // Command direction FW M2CM9S
        [3].4   // VMCC M2 Speed zone 5 Drive Fault * 2CM05S
        [3].10   // VMCC M2 Speed zone 11 Drive Fault 2CM11S
        [32].1   // PANEL KD-CS1N Knurl knocker Move OUT South Selector Sw.
        [3].5   // VMCC M2 Speed zone 6 Drive Fault * 2CM06S
        [4].10   // VMCC M2 Speed zone 11 Drive Fault 2CM11N
        [76].5   // PANEL KD-CS1S Knurl knocker Move DOWN South Selector Sw.
        [24].13   // RELIANCE CAPPING SYSTEM Adapter Power ON
        [72].11   // BENCHBOARD Trim knocker #3 South Auto mode
        [3].11   // VMCC M2 Speed zone 12 Drive Fault * 2CM12S
        [72].13   // BENCHBOARD Trim knocker #4 North Auto mode
        [123].2   // MB -->> M2 Reliance Crossbreak In progres
        [123].1   // MB -->> M2 Crossbreak In progress Front end
        [33].6   // PANEL KD-CS1N Trim deck North Outer Limit Sw.
        [17].1   // VMCC TD Drive Contactor Energized
        [18].0   // VMCC TD Trim knocker Drive fault
        [2].12   // VMCC M2 Drive Comm Module Power On
        [18].4   // VMCC TD Trim deck Alarm lamp
        [24].11   // RELIANCE CAPPING SYSTEM
        [2].2   // VMCC M2 DC Input Power ON
        [101].11   // Local control 3 M2CM8S
        [101].7   // Drive has a fault M2CM8S
        [105].3   // Actual direction FWD M2CM9S
        [101].9   // Local control 1 M2CM8S
        [103].10   // Local control 2 M2CM8N
        [101].15   // Speed reference 4 M2CM8S
        [111].14   // Speed reference 3 M2CM10N
        [105].7   // Drive has a fault M2CM9S
        [107].10   // Local control 2 M2CM9N
        [111].0   // Drive ready M2CM10N
        [100]   // RACK 14 INPUT UPDATES
        [111].15   // Speed reference 4 M2CM10N
        [111].2   // Command direction FW M2CM10N
        [111].3   // Actual direction FWD M2CM10N
        [111].6   // Drive has an alarm M2CM10N
        [113].12   // Speed reference 1 M2CM11S
        [113].13   // Speed reference 2 M2CM11S
        [113].14   // Speed reference 3 M2CM11S
        [113].15   // Speed reference 4 M2CM11S
        [113].2   // Command direction FW M2CM11S
        [115].15   // Speed reference 4 M2CM11N
        [2].1   // VMCC M2 Drive Contactor Energized
        [2].11   // VMCC M2 Panel Overtemp Alarm
        [107].0   // Drive ready M2CM9N
        [2].6   // VMCC M2 DC Power Supply #1 ON
        [2].7   // VMCC M2 DC Power Supply #2 ON
        [65].15   // PANEL TD-CS3S SPARE
        [68].12   // PANEL TD-CS2S SPARE
        [68].13   // PANEL TD-CS2S SPARE
        [68].14   // PANEL TD-CS2S SPARE
        [68].15   // PANEL TD-CS2S SPARE
        [107].12   // Speed reference 1 M2CM9N
        [107].13   // Speed reference 2 M2CM9N
        [1].8   // Rockwell Run out Speed up signal M2CM10
        [1].9   // Rockwell Run out Speed up signal M2CM11
        [113].3   // Actual direction FWD M2CM11S
        [123].4   // MB -->> M2 Eclipse Mode Operation On
        [115].2   // Command direction FW M2CM11N
        [115].3   // Actual direction FWD M2CM11N
        [115].6   // Drive has an alarm M2CM11N
        [115].7   // Drive has a fault M2CM11N
        [69].14   // PANEL TD-CS2S SPARE
        [103].12   // Speed reference 1 M2CM8N
        [101].3   // Actual direction FWD M2CM8S
        [107].14   // Speed reference 3 M2CM9N
        [117].10   // Local control 2 M2CM12S
        [123].10   // MB -->> M2 SPARE
        [103].9   // Local control 1 M2CM8N
        [103].13   // Speed reference 2 M2CM8N
        [72].4   // BENCHBOARD Trim knocker #2 North Up Selector Sw.
        [73].1   // BENCHBOARD Knocker #5 North Auto mode
        [107].15   // Speed reference 4 M2CM9N
        [72].15   // BENCHBOARD Trim knocker #4 South Auto mode
        [113].6   // Drive has an alarm M2CM11S
        [1].1   // Rockwell Run out Speed up signal M2CM3
        [33].7   // PANEL KD-CS1N Trim deck North Inner Limit Sw.
        [1].2   // Rockwell Run out Speed up signal M2CM4
        [115].10   // Local control 2 M2CM11N
        [69].15   // PANEL TD-CS2S SPARE
        [117].11   // Local control 3 M2CM12S
        [117].12   // Speed reference 1 M2CM12S
        [73].12   // BENCHBOARD Drop No. 1 Crusher
        [73].13   // BENCHBOARD Adapter Power ON
        [115].11   // Local control 3 M2CM11N
        [32].7   // PANEL KD-CS1N Knurl knocker Move OUT North Selector Sw.
        [36].0   // PANEL TD-CS1N Trim knocker 1 Move IN South Selector Sw.
        [36].15   // PANEL TD-CS1N Eclipse Hold Down Wheels Up Sel. Sw.
        [107].2   // Command direction FW M2CM9N
        [1].3   // Rockwell Run out Speed up signal M2CM5
        [107].3   // Actual direction FWD M2CM9N
        [109].12   // Speed reference 1 M2CM10S
        [109].13   // Speed reference 2 M2CM10S
        [1].4   // Rockwell Run out Speed up signal M2CM6
        [125].0   // ROCKWELL CAPPER Input for crossbreak in progress
